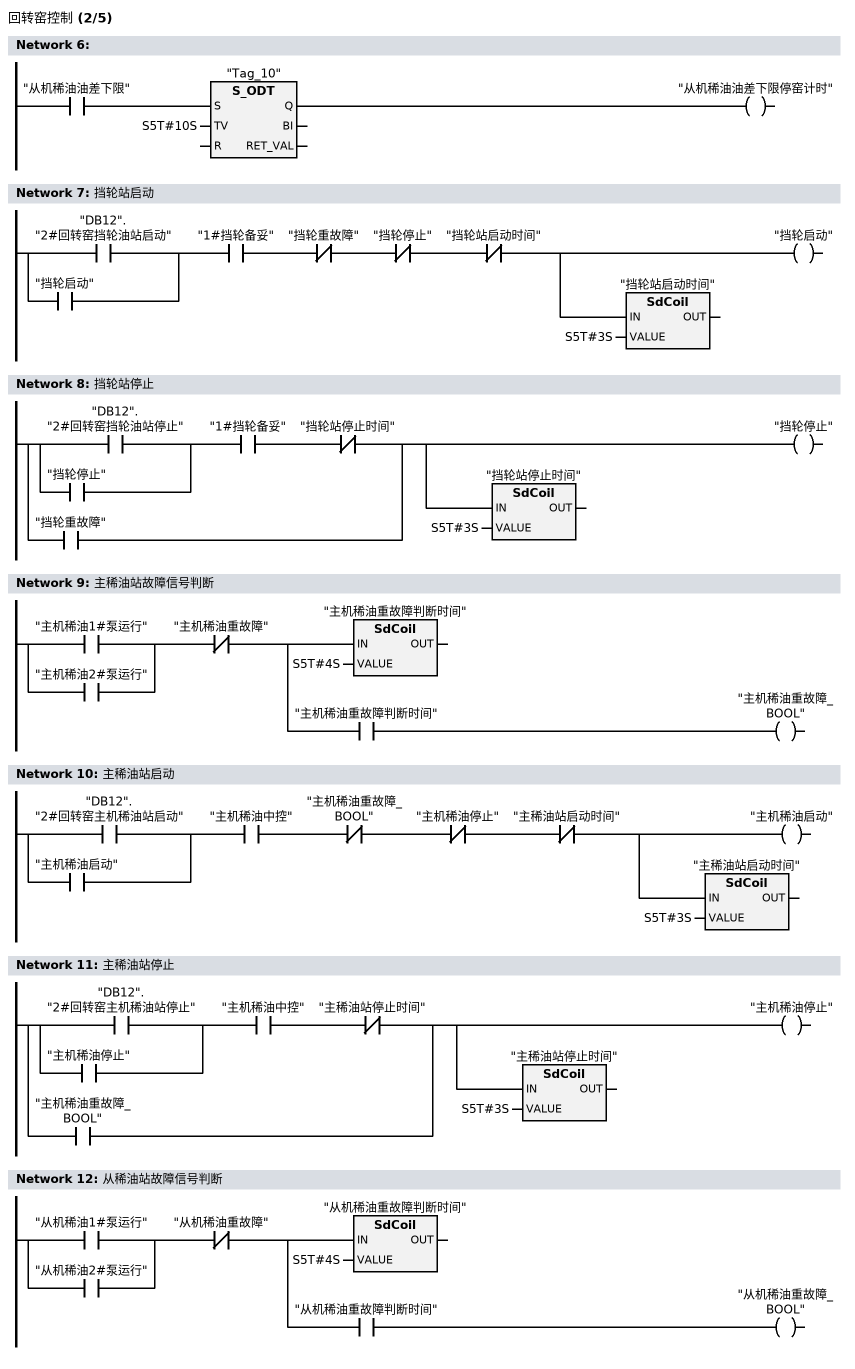
   RUNG wire#powerrail
      Contact( "从机稀油油差下限" )
      S_ODT(T_NO := "Tag_10", TV := S5T#10S, R :=, BI =>, RET_VAL =>)
      Coil( "从机稀油油差下限停窑计时" )
   END_RUNG
   // the same network as SCL:
   #_s5time1 := S_ODT(T_NO := "Tag_10", TV := S5T#10S, S := "从机稀油油差下限", Q => #_w1);
   "从机稀油油差下限停窑计时" := #_w1;
END_REGION

REGION Network 7: 挡轮站启动
   // no SCL statement known for SdCoil: written as a call
   "挡轮启动" := ("DB12"."2#回转窑挡轮油站启动" OR "挡轮启动") AND "1#挡轮备妥" AND NOT "挡轮重故障" AND NOT "挡轮停止" AND NOT "挡轮站启动时间";
   SdCoil(in := "挡轮启动", value := S5T#3S, operand := "挡轮站启动时间");
END_REGION

REGION Network 8: 挡轮站停止
   // no SCL statement known for SdCoil: written as a call
   "挡轮停止" := (("DB12"."2#回转窑挡轮油站停止" OR "挡轮停止") AND "1#挡轮备妥" AND NOT "挡轮站停止时间") OR "挡轮重故障";
   SdCoil(in := "挡轮停止", value := S5T#3S, operand := "挡轮站停止时间");
END_REGION

REGION Network 9: 主稀油站故障信号判断
   // no SCL statement known for SdCoil: written as a call
   #_w1 := ("主机稀油1#泵运行" OR "主机稀油2#泵运行") AND NOT "主机稀油重故障";
   SdCoil(in := #_w1, value := S5T#4S, operand := "主机稀油重故障判断时间");
   "主机稀油重故障_BOOL" := #_w1 AND "主机稀油重故障判断时间";
END_REGION

REGION Network 10: 主稀油站启动
   // no SCL statement known for SdCoil: written as a call
   "主机稀油启动" := ("DB12"."2#回转窑主机稀油站启动" OR "主机稀油启动") AND "主机稀油中控" AND NOT "主机稀油重故障_BOOL" AND NOT "主机稀油停止" AND NOT "主稀油站启动时间";
   SdCoil(in := "主机稀油启动", value := S5T#3S, operand := "主稀油站启动时间");
END_REGION

REGION Network 11: 主稀油站停止
   // no SCL statement known for SdCoil: written as a call
   "主机稀油停止" := (("DB12"."2#回转窑主机稀油站停止" OR "主机稀油停止") AND "主机稀油中控" AND NOT "主稀油站停止时间") OR "主机稀油重故障_BOOL";
   SdCoil(in := "主机稀油停止", value := S5T#3S, operand := "主稀油站停止时间");
END_REGION

REGION Network 12: 从稀油站故障信号判断
   // no SCL statement known for SdCoil: written as a call
   #_w1 := ("从机稀油1#泵运行" OR "从机稀油2#泵运行") AND NOT "从机稀油重故障";
   SdCoil(in := #_w1, value := S5T#4S, operand := "从机稀油重故障判断时间");
   "从机稀油重故障_BOOL" := #_w1 AND "从机稀油重故障判断时间";
END_REGION

REGION Network 13: 从稀油站启动
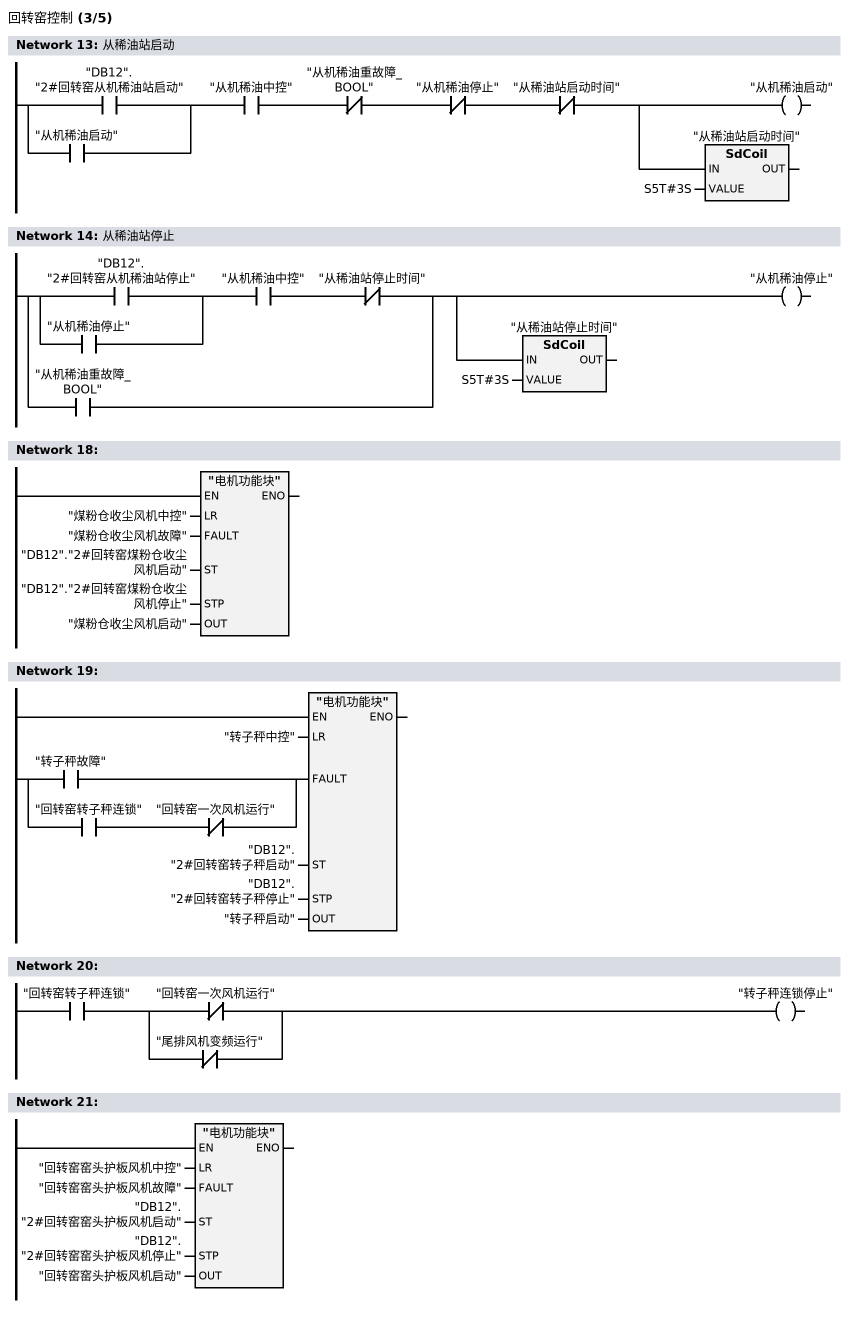
   // no SCL statement known for SdCoil: written as a call
   "从机稀油启动" := ("DB12"."2#回转窑从机稀油站启动" OR "从机稀油启动") AND "从机稀油中控" AND NOT "从机稀油重故障_BOOL" AND NOT "从机稀油停止" AND NOT "从稀油站启动时间";
   SdCoil(in := "从机稀油启动", value := S5T#3S, operand := "从稀油站启动时间");
END_REGION

REGION Network 14: 从稀油站停止
   // no SCL statement known for SdCoil: written as a call
   "从机稀油停止" := (("DB12"."2#回转窑从机稀油站停止" OR "从机稀油停止") AND "从机稀油中控" AND NOT "从稀油站停止时间") OR "从机稀油重故障_BOOL";
   SdCoil(in := "从机稀油停止", value := S5T#3S, operand := "从稀油站停止时间");
END_REGION

REGION Network 18
   RUNG wire#powerrail
      "电机功能块"(LR := "煤粉仓收尘风机中控", FAULT := "煤粉仓收尘风机故障", ST := "DB12"."2#回转窑煤粉仓收尘风机启动", STP := "DB12"."2#回转窑煤粉仓收尘风机停止", OUT := "煤粉仓收尘风机启动")
   END_RUNG
   // the same network as SCL:
   "电机功能块"(LR := "煤粉仓收尘风机中控",
           FAULT := "煤粉仓收尘风机故障",
           ST := "DB12"."2#回转窑煤粉仓收尘风机启动",
           STP := "DB12"."2#回转窑煤粉仓收尘风机停止",
           OUT := "煤粉仓收尘风机启动");
END_REGION

REGION Network 19
   RUNG wire#powerrail
      "电机功能块"(FAULT := wire#w1, LR := "转子秤中控", ST := "DB12"."2#回转窑转子秤启动", STP := "DB12"."2#回转窑转子秤停止", OUT := "转子秤启动")
   END_RUNG
   RUNG wire#powerrail
      Contact( "转子秤故障" )
   END_RUNG wire#w1
   RUNG wire#powerrail
      Contact( "回转窑转子秤连锁" )
      I_Contact( "回转窑一次风机运行" )
   END_RUNG wire#w1
   // the same network as SCL:
   "电机功能块"(LR := "转子秤中控",
           FAULT := "转子秤故障" OR ("回转窑转子秤连锁" AND NOT "回转窑一次风机运行"),
           ST := "DB12"."2#回转窑转子秤启动",
           STP := "DB12"."2#回转窑转子秤停止",
           OUT := "转子秤启动");
END_REGION

REGION Network 20
   RUNG wire#powerrail
      Contact( "回转窑转子秤连锁" )
      wire#w1
      I_Contact( "回转窑一次风机运行" )
      wire#w2
      Coil( "转子秤连锁停止" )
   END_RUNG
   RUNG wire#w1
      I_Contact( "尾排风机变频运行" )
   END_RUNG wire#w2
   // the same network as SCL:
   "转子秤连锁停止" := "回转窑转子秤连锁" AND (NOT "回转窑一次风机运行" OR NOT "尾排风机变频运行");
END_REGION

REGION Network 21
   RUNG wire#powerrail
      "电机功能块"(LR := "回转窑窑头护板风机中控", FAULT := "回转窑窑头护板风机故障", ST := "DB12"."2#回转窑窑头护板风机启动", STP := "DB12"."2#回转窑窑头护板风机停止", OUT := "回转窑窑头护板风机启动")
   END_RUNG
   // the same network as SCL:
   "电机功能块"(LR := "回转窑窑头护板风机中控",
           FAULT := "回转窑窑头护板风机故障",
           ST := "DB12"."2#回转窑窑头护板风机启动",
           STP := "DB12"."2#回转窑窑头护板风机停止",
           OUT := "回转窑窑头护板风机启动");
END_REGION

REGION Network 22
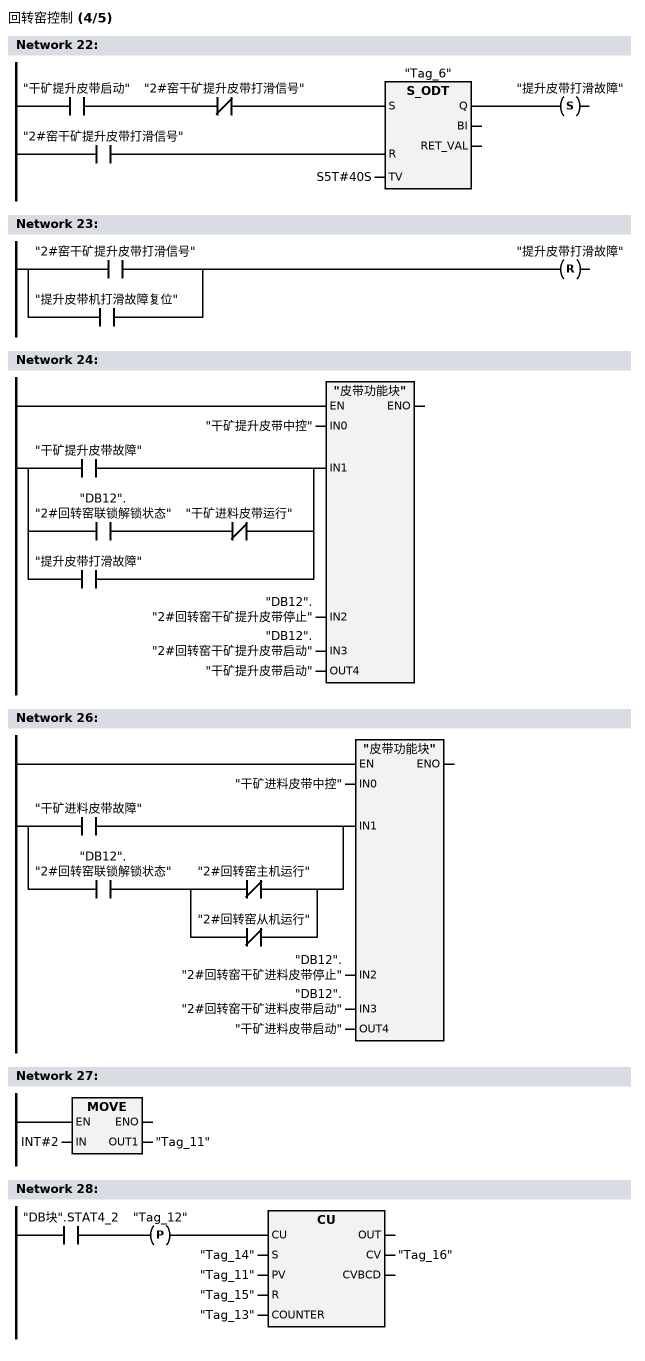
   RUNG wire#powerrail
      Contact( "干矿提升皮带启动" )
      I_Contact( "2#窑干矿提升皮带打滑信号" )
      S_ODT(T_NO := "Tag_6", R := wire#w1, TV := S5T#40S, BI =>, RET_VAL =>)
      S_Coil( "提升皮带打滑故障" )
   END_RUNG
   RUNG wire#powerrail
      Contact( "2#窑干矿提升皮带打滑信号" )
   END_RUNG wire#w1
   // the same network as SCL:
   #_s5time1 := S_ODT(T_NO := "Tag_6",
                      S := "干矿提升皮带启动" AND NOT "2#窑干矿提升皮带打滑信号",
                      R := "2#窑干矿提升皮带打滑信号",
                      TV := S5T#40S,
                      Q => #_w1);
   IF #_w1 THEN "提升皮带打滑故障" := TRUE; END_IF;
END_REGION

REGION Network 23
   RUNG wire#powerrail
      Contact( "2#窑干矿提升皮带打滑信号" )
      wire#w1
      R_Coil( "提升皮带打滑故障" )
   END_RUNG
   RUNG wire#powerrail
      Contact( "提升皮带机打滑故障复位" )
   END_RUNG wire#w1
   // the same network as SCL:
   IF "2#窑干矿提升皮带打滑信号" OR "提升皮带机打滑故障复位" THEN "提升皮带打滑故障" := FALSE; END_IF;
END_REGION

REGION Network 24
   RUNG wire#powerrail
      "皮带功能块"(IN1 := wire#w1, IN0 := "干矿提升皮带中控", IN2 := "DB12"."2#回转窑干矿提升皮带停止", IN3 := "DB12"."2#回转窑干矿提升皮带启动", OUT4 := "干矿提升皮带启动")
   END_RUNG
   RUNG wire#powerrail
      Contact( "干矿提升皮带故障" )
   END_RUNG wire#w1
   RUNG wire#powerrail
      Contact( "DB12"."2#回转窑联锁解锁状态" )
      I_Contact( "干矿进料皮带运行" )
   END_RUNG wire#w1
   RUNG wire#powerrail
      Contact( "提升皮带打滑故障" )
   END_RUNG wire#w1
   // the same network as SCL:
   "皮带功能块"(IN0 := "干矿提升皮带中控",
           IN1 := "干矿提升皮带故障" OR ("DB12"."2#回转窑联锁解锁状态" AND NOT "干矿进料皮带运行") OR "提升皮带打滑故障",
           IN2 := "DB12"."2#回转窑干矿提升皮带停止",
           IN3 := "DB12"."2#回转窑干矿提升皮带启动",
           OUT4 := "干矿提升皮带启动");
END_REGION

REGION Network 26
   RUNG wire#powerrail
      "皮带功能块"(IN1 := wire#w2, IN0 := "干矿进料皮带中控", IN2 := "DB12"."2#回转窑干矿进料皮带停止", IN3 := "DB12"."2#回转窑干矿进料皮带启动", OUT4 := "干矿进料皮带启动")
   END_RUNG
   RUNG wire#powerrail
      Contact( "干矿进料皮带故障" )
   END_RUNG wire#w2
   RUNG wire#powerrail
      Contact( "DB12"."2#回转窑联锁解锁状态" )
      wire#w1
      I_Contact( "2#回转窑主机运行" )
   END_RUNG wire#w2
   RUNG wire#w1
      I_Contact( "2#回转窑从机运行" )
   END_RUNG wire#w2
   // the same network as SCL:
   "皮带功能块"(IN0 := "干矿进料皮带中控",
           IN1 := "干矿进料皮带故障" OR ("DB12"."2#回转窑联锁解锁状态" AND (NOT "2#回转窑主机运行" OR NOT "2#回转窑从机运行")),
           IN2 := "DB12"."2#回转窑干矿进料皮带停止",
           IN3 := "DB12"."2#回转窑干矿进料皮带启动",
           OUT4 := "干矿进料皮带启动");
END_REGION

REGION Network 27
   RUNG wire#powerrail
      { S7_GenerateENO := "TRUE" } Move(in := INT#2, out1 => "Tag_11")
   END_RUNG
   // the same network as SCL:
   "Tag_11" := INT#2;
END_REGION

REGION Network 28
   // no SCL statement known for Cu: written as a call
   #_w1 := "DB块".STAT4_2 AND NOT "Tag_12";   // rising edge
   "Tag_12" := "DB块".STAT4_2;
   Cu(cu := #_w1, s := "Tag_14", pv := "Tag_11", r := "Tag_15", "counter" := "Tag_13", cv => "Tag_16");
END_REGION

REGION Network 29
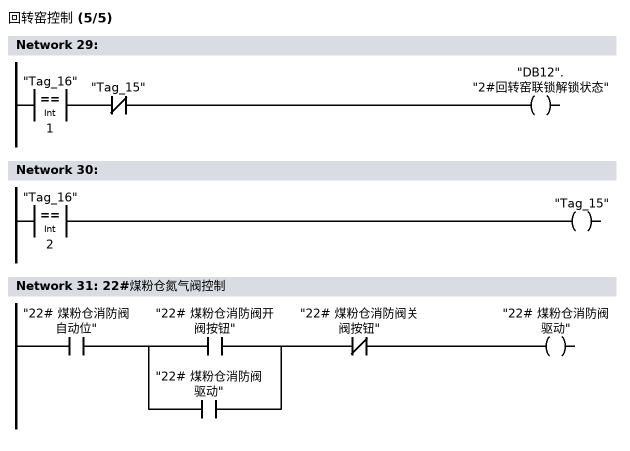
   RUNG wire#powerrail
      { S7_Templates := "SrcType := Int" } EQ_Contact(in1 := "Tag_16", in2 := 1)
      I_Contact( "Tag_15" )
      Coil( "DB12"."2#回转窑联锁解锁状态" )
   END_RUNG
   // the same network as SCL:
   "DB12"."2#回转窑联锁解锁状态" := ("Tag_16" = 1) AND NOT "Tag_15";
END_REGION

REGION Network 30
   RUNG wire#powerrail
      { S7_Templates := "SrcType := Int" } EQ_Contact(in1 := "Tag_16", in2 := 2)
      Coil( "Tag_15" )
   END_RUNG
   // the same network as SCL:
   "Tag_15" := "Tag_16" = 2;
END_REGION

REGION Network 31: 22#煤粉仓氮气阀控制
   RUNG wire#powerrail
      Contact( "22# 煤粉仓消防阀自动位" )
      wire#w1
      Contact( "22# 煤粉仓消防阀开阀按钮" )
      wire#w2
      I_Contact( "22# 煤粉仓消防阀关阀按钮" )
      Coil( "22# 煤粉仓消防阀驱动" )
   END_RUNG
   RUNG wire#w1
      Contact( "22# 煤粉仓消防阀驱动" )
   END_RUNG wire#w2
   // the same network as SCL:
   "22# 煤粉仓消防阀驱动" := "22# 煤粉仓消防阀自动位" AND ("22# 煤粉仓消防阀开阀按钮" OR "22# 煤粉仓消防阀驱动") AND NOT "22# 煤粉仓消防阀关阀按钮";
END_REGION
END_FUNCTION

FUNCTION "回转窑模拟量反馈" : Void   // FC12, LAD
{ S7_Optimized_Access := 'FALSE' }
VERSION : 0.1
   VAR_TEMP   // added for the SCL form of the ladder/FBD networks
      _w1 : Bool;
      _s5time1 : S5Time;
   END_VAR
BEGIN

REGION Network 1
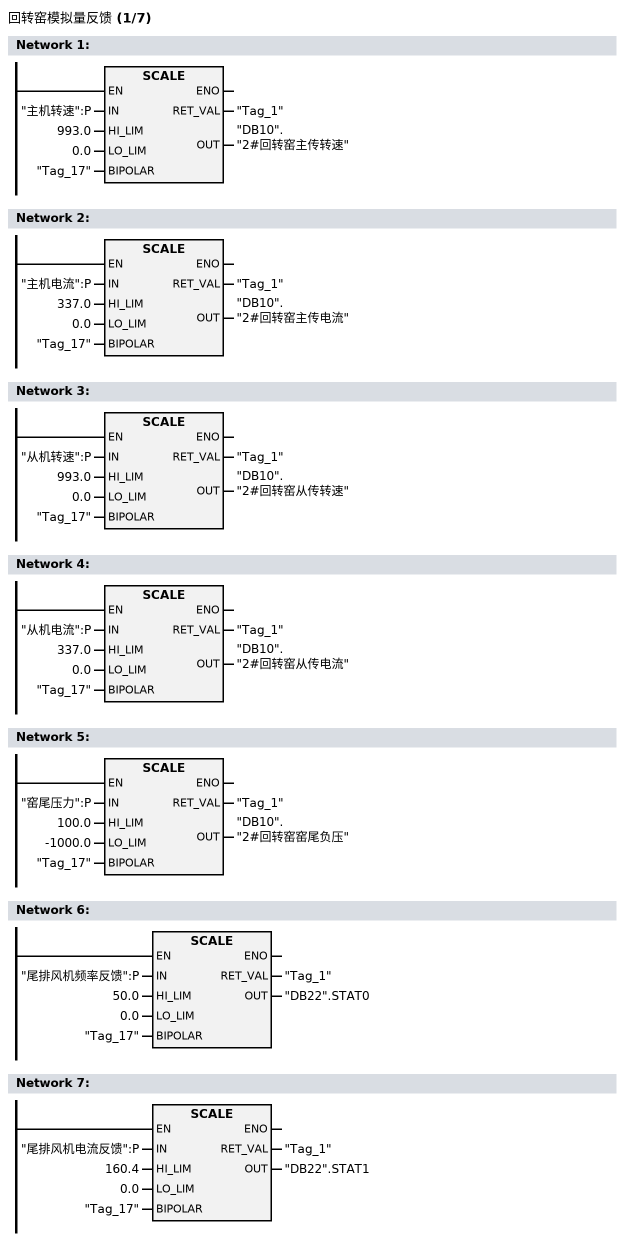
   "Tag_1" := SCALE(IN := "主机转速":P,
                    HI_LIM := 993.0,
                    LO_LIM := 0.0,
                    BIPOLAR := "Tag_17",
                    OUT => "DB10"."2#回转窑主传转速");
END_REGION

REGION Network 2
   "Tag_1" := SCALE(IN := "主机电流":P,
                    HI_LIM := 337.0,
                    LO_LIM := 0.0,
                    BIPOLAR := "Tag_17",
                    OUT => "DB10"."2#回转窑主传电流");
END_REGION

REGION Network 3
   "Tag_1" := SCALE(IN := "从机转速":P,
                    HI_LIM := 993.0,
                    LO_LIM := 0.0,
                    BIPOLAR := "Tag_17",
                    OUT => "DB10"."2#回转窑从传转速");
END_REGION

REGION Network 4
   "Tag_1" := SCALE(IN := "从机电流":P,
                    HI_LIM := 337.0,
                    LO_LIM := 0.0,
                    BIPOLAR := "Tag_17",
                    OUT => "DB10"."2#回转窑从传电流");
END_REGION

REGION Network 5
   "Tag_1" := SCALE(IN := "窑尾压力":P,
                    HI_LIM := 100.0,
                    LO_LIM := -1000.0,
                    BIPOLAR := "Tag_17",
                    OUT => "DB10"."2#回转窑窑尾负压");
END_REGION

REGION Network 6
   "Tag_1" := SCALE(IN := "尾排风机频率反馈":P, HI_LIM := 50.0, LO_LIM := 0.0, BIPOLAR := "Tag_17", OUT => "DB22".STAT0);
END_REGION

REGION Network 7
   "Tag_1" := SCALE(IN := "尾排风机电流反馈":P,
                    HI_LIM := 160.4,
                    LO_LIM := 0.0,
                    BIPOLAR := "Tag_17",
                    OUT => "DB22".STAT1);
END_REGION

REGION Network 8
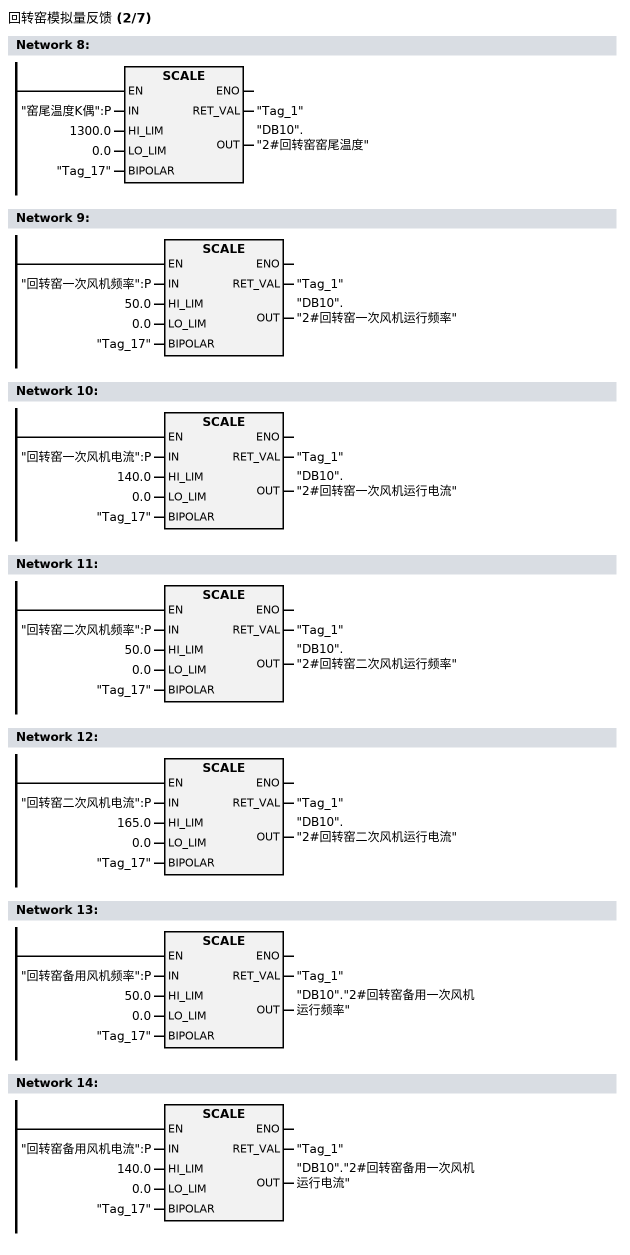
   "Tag_1" := SCALE(IN := "窑尾温度K偶":P,
                    HI_LIM := 1300.0,
                    LO_LIM := 0.0,
                    BIPOLAR := "Tag_17",
                    OUT => "DB10"."2#回转窑窑尾温度");
END_REGION

REGION Network 9
   "Tag_1" := SCALE(IN := "回转窑一次风机频率":P,
                    HI_LIM := 50.0,
                    LO_LIM := 0.0,
                    BIPOLAR := "Tag_17",
                    OUT => "DB10"."2#回转窑一次风机运行频率");
END_REGION

REGION Network 10
   "Tag_1" := SCALE(IN := "回转窑一次风机电流":P,
                    HI_LIM := 140.0,
                    LO_LIM := 0.0,
                    BIPOLAR := "Tag_17",
                    OUT => "DB10"."2#回转窑一次风机运行电流");
END_REGION

REGION Network 11
   "Tag_1" := SCALE(IN := "回转窑二次风机频率":P,
                    HI_LIM := 50.0,
                    LO_LIM := 0.0,
                    BIPOLAR := "Tag_17",
                    OUT => "DB10"."2#回转窑二次风机运行频率");
END_REGION

REGION Network 12
   "Tag_1" := SCALE(IN := "回转窑二次风机电流":P,
                    HI_LIM := 165.0,
                    LO_LIM := 0.0,
                    BIPOLAR := "Tag_17",
                    OUT => "DB10"."2#回转窑二次风机运行电流");
END_REGION

REGION Network 13
   "Tag_1" := SCALE(IN := "回转窑备用风机频率":P,
                    HI_LIM := 50.0,
                    LO_LIM := 0.0,
                    BIPOLAR := "Tag_17",
                    OUT => "DB10"."2#回转窑备用一次风机运行频率");
END_REGION

REGION Network 14
   "Tag_1" := SCALE(IN := "回转窑备用风机电流":P,
                    HI_LIM := 140.0,
                    LO_LIM := 0.0,
                    BIPOLAR := "Tag_17",
                    OUT => "DB10"."2#回转窑备用一次风机运行电流");
END_REGION

REGION Network 15
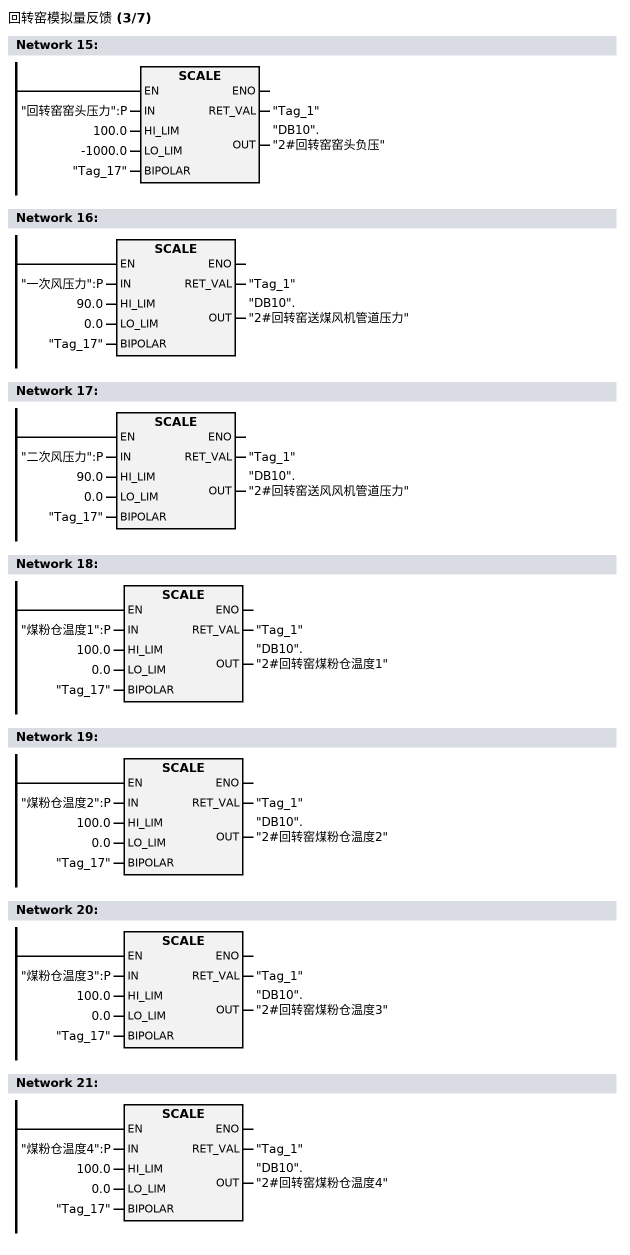
   "Tag_1" := SCALE(IN := "回转窑窑头压力":P,
                    HI_LIM := 100.0,
                    LO_LIM := -1000.0,
                    BIPOLAR := "Tag_17",
                    OUT => "DB10"."2#回转窑窑头负压");
END_REGION

REGION Network 16
   "Tag_1" := SCALE(IN := "一次风压力":P,
                    HI_LIM := 90.0,
                    LO_LIM := 0.0,
                    BIPOLAR := "Tag_17",
                    OUT => "DB10"."2#回转窑送煤风机管道压力");
END_REGION

REGION Network 17
   "Tag_1" := SCALE(IN := "二次风压力":P,
                    HI_LIM := 90.0,
                    LO_LIM := 0.0,
                    BIPOLAR := "Tag_17",
                    OUT => "DB10"."2#回转窑送风风机管道压力");
END_REGION

REGION Network 18
   "Tag_1" := SCALE(IN := "煤粉仓温度1":P,
                    HI_LIM := 100.0,
                    LO_LIM := 0.0,
                    BIPOLAR := "Tag_17",
                    OUT => "DB10"."2#回转窑煤粉仓温度1");
END_REGION

REGION Network 19
   "Tag_1" := SCALE(IN := "煤粉仓温度2":P,
                    HI_LIM := 100.0,
                    LO_LIM := 0.0,
                    BIPOLAR := "Tag_17",
                    OUT => "DB10"."2#回转窑煤粉仓温度2");
END_REGION

REGION Network 20
   "Tag_1" := SCALE(IN := "煤粉仓温度3":P,
                    HI_LIM := 100.0,
                    LO_LIM := 0.0,
                    BIPOLAR := "Tag_17",
                    OUT => "DB10"."2#回转窑煤粉仓温度3");
END_REGION

REGION Network 21
   "Tag_1" := SCALE(IN := "煤粉仓温度4":P,
                    HI_LIM := 100.0,
                    LO_LIM := 0.0,
                    BIPOLAR := "Tag_17",
                    OUT => "DB10"."2#回转窑煤粉仓温度4");
END_REGION

REGION Network 22
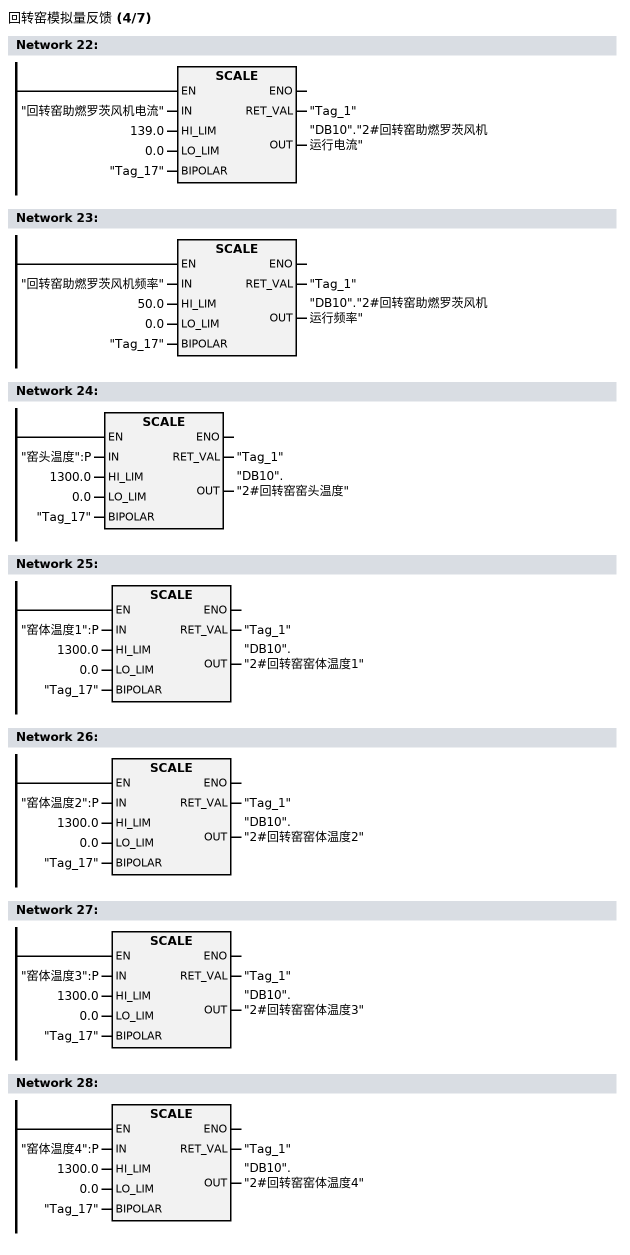
   "Tag_1" := SCALE(IN := "回转窑助燃罗茨风机电流",
                    HI_LIM := 139.0,
                    LO_LIM := 0.0,
                    BIPOLAR := "Tag_17",
                    OUT => "DB10"."2#回转窑助燃罗茨风机运行电流");
END_REGION

REGION Network 23
   "Tag_1" := SCALE(IN := "回转窑助燃罗茨风机频率",
                    HI_LIM := 50.0,
                    LO_LIM := 0.0,
                    BIPOLAR := "Tag_17",
                    OUT => "DB10"."2#回转窑助燃罗茨风机运行频率");
END_REGION

REGION Network 24
   "Tag_1" := SCALE(IN := "窑头温度":P,
                    HI_LIM := 1300.0,
                    LO_LIM := 0.0,
                    BIPOLAR := "Tag_17",
                    OUT => "DB10"."2#回转窑窑头温度");
END_REGION

REGION Network 25
   "Tag_1" := SCALE(IN := "窑体温度1":P,
                    HI_LIM := 1300.0,
                    LO_LIM := 0.0,
                    BIPOLAR := "Tag_17",
                    OUT => "DB10"."2#回转窑窑体温度1");
END_REGION

REGION Network 26
   "Tag_1" := SCALE(IN := "窑体温度2":P,
                    HI_LIM := 1300.0,
                    LO_LIM := 0.0,
                    BIPOLAR := "Tag_17",
                    OUT => "DB10"."2#回转窑窑体温度2");
END_REGION

REGION Network 27
   "Tag_1" := SCALE(IN := "窑体温度3":P,
                    HI_LIM := 1300.0,
                    LO_LIM := 0.0,
                    BIPOLAR := "Tag_17",
                    OUT => "DB10"."2#回转窑窑体温度3");
END_REGION

REGION Network 28
   "Tag_1" := SCALE(IN := "窑体温度4":P,
                    HI_LIM := 1300.0,
                    LO_LIM := 0.0,
                    BIPOLAR := "Tag_17",
                    OUT => "DB10"."2#回转窑窑体温度4");
END_REGION

REGION Network 29
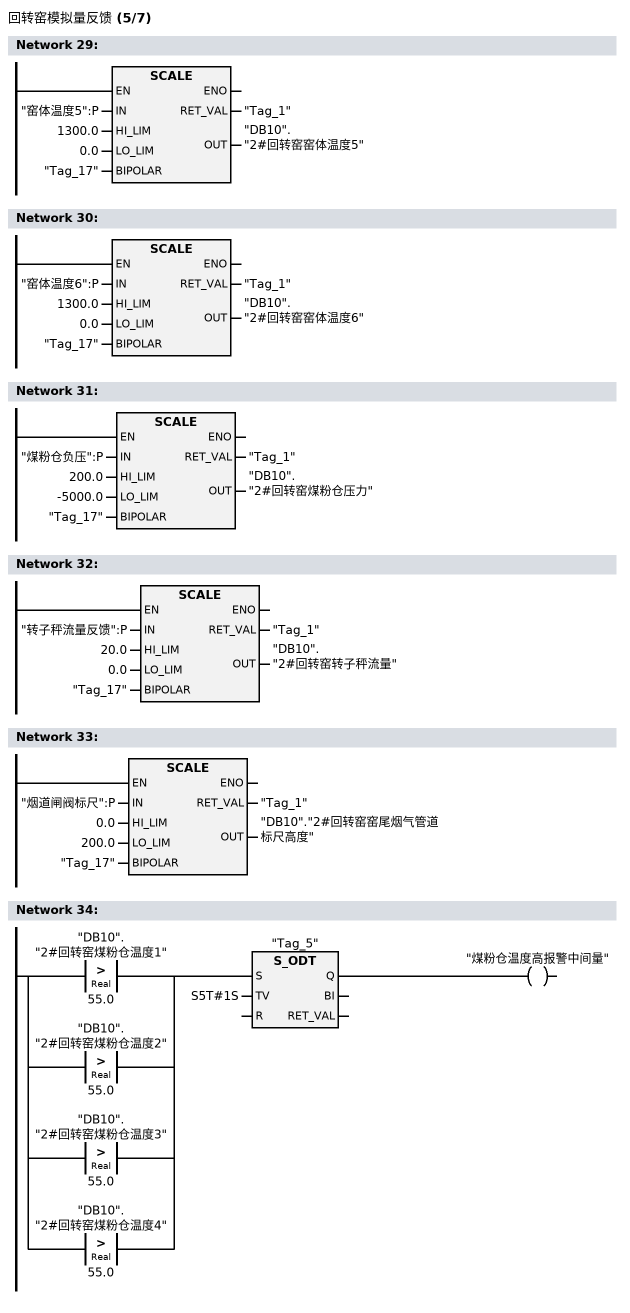
   "Tag_1" := SCALE(IN := "窑体温度5":P,
                    HI_LIM := 1300.0,
                    LO_LIM := 0.0,
                    BIPOLAR := "Tag_17",
                    OUT => "DB10"."2#回转窑窑体温度5");
END_REGION

REGION Network 30
   "Tag_1" := SCALE(IN := "窑体温度6":P,
                    HI_LIM := 1300.0,
                    LO_LIM := 0.0,
                    BIPOLAR := "Tag_17",
                    OUT => "DB10"."2#回转窑窑体温度6");
END_REGION

REGION Network 31
   "Tag_1" := SCALE(IN := "煤粉仓负压":P,
                    HI_LIM := 200.0,
                    LO_LIM := -5000.0,
                    BIPOLAR := "Tag_17",
                    OUT => "DB10"."2#回转窑煤粉仓压力");
END_REGION

REGION Network 32
   "Tag_1" := SCALE(IN := "转子秤流量反馈":P,
                    HI_LIM := 20.0,
                    LO_LIM := 0.0,
                    BIPOLAR := "Tag_17",
                    OUT => "DB10"."2#回转窑转子秤流量");
END_REGION

REGION Network 33
   "Tag_1" := SCALE(IN := "烟道闸阀标尺":P,
                    HI_LIM := 0.0,
                    LO_LIM := 200.0,
                    BIPOLAR := "Tag_17",
                    OUT => "DB10"."2#回转窑窑尾烟气管道标尺高度");
END_REGION

REGION Network 34
   RUNG wire#powerrail
      { S7_Templates := "SrcType := Real" } GT_Contact(in1 := "DB10"."2#回转窑煤粉仓温度1", in2 := 55.0)
      wire#w1
      S_ODT(T_NO := "Tag_5", TV := S5T#1S, R :=, BI =>, RET_VAL =>)
      Coil( "煤粉仓温度高报警中间量" )
   END_RUNG
   RUNG wire#powerrail
      { S7_Templates := "SrcType := Real" } GT_Contact(in1 := "DB10"."2#回转窑煤粉仓温度2", in2 := 55.0)
   END_RUNG wire#w1
   RUNG wire#powerrail
      { S7_Templates := "SrcType := Real" } GT_Contact(in1 := "DB10"."2#回转窑煤粉仓温度3", in2 := 55.0)
   END_RUNG wire#w1
   RUNG wire#powerrail
      { S7_Templates := "SrcType := Real" } GT_Contact(in1 := "DB10"."2#回转窑煤粉仓温度4", in2 := 55.0)
   END_RUNG wire#w1
   // the same network as SCL:
   #_s5time1 := S_ODT(T_NO := "Tag_5",
                      S := ("DB10"."2#回转窑煤粉仓温度1" > 55.0) OR ("DB10"."2#回转窑煤粉仓温度2" > 55.0) OR ("DB10"."2#回转窑煤粉仓温度3" > 55.0) OR ("DB10"."2#回转窑煤粉仓温度4" > 55.0),
                      TV := S5T#1S,
                      Q => #_w1);
   "煤粉仓温度高报警中间量" := #_w1;
END_REGION

REGION Network 35
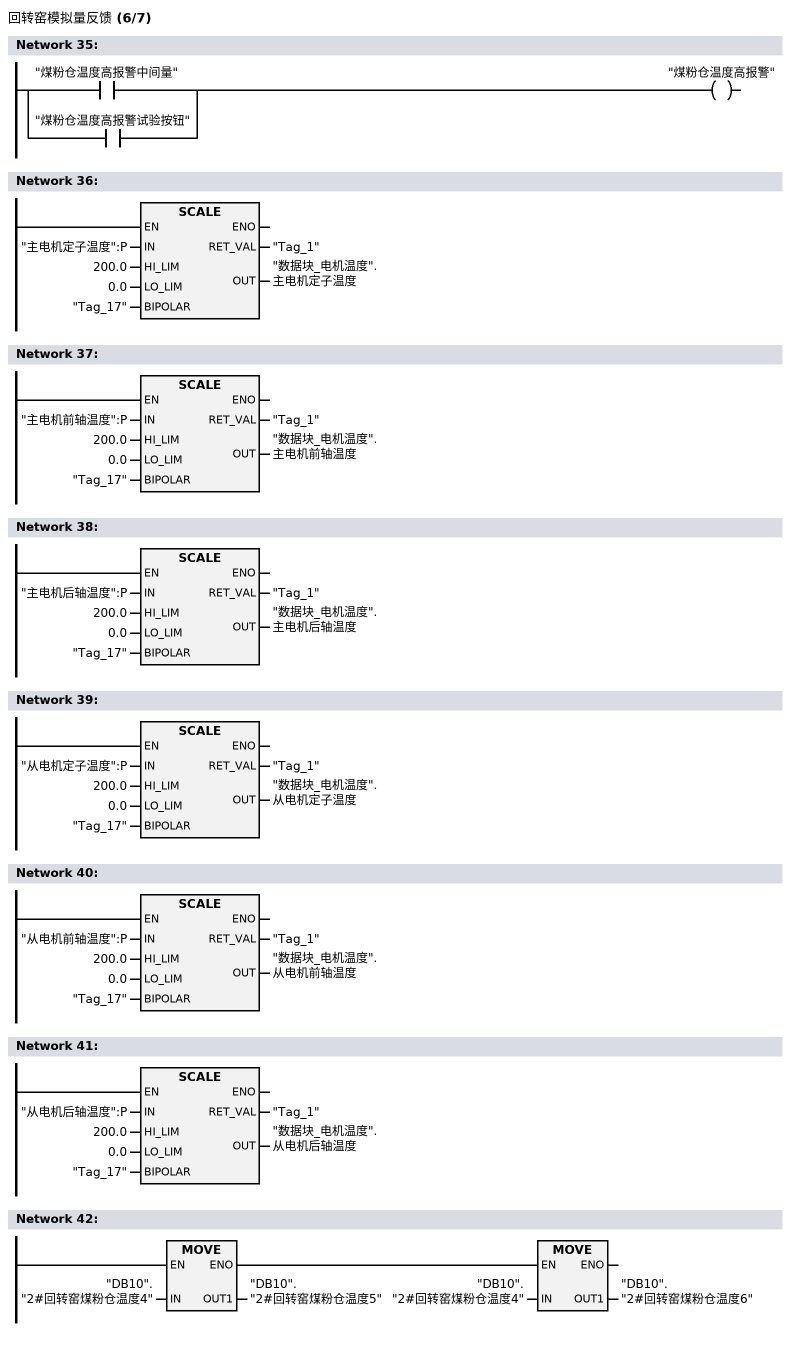
   RUNG wire#powerrail
      Contact( "煤粉仓温度高报警中间量" )
      wire#w1
      Coil( "煤粉仓温度高报警" )
   END_RUNG
   RUNG wire#powerrail
      Contact( "煤粉仓温度高报警试验按钮" )
   END_RUNG wire#w1
   // the same network as SCL:
   "煤粉仓温度高报警" := "煤粉仓温度高报警中间量" OR "煤粉仓温度高报警试验按钮";
END_REGION

REGION Network 36
   "Tag_1" := SCALE(IN := "主电机定子温度":P,
                    HI_LIM := 200.0,
                    LO_LIM := 0.0,
                    BIPOLAR := "Tag_17",
                    OUT => "数据块_电机温度".主电机定子温度);
END_REGION

REGION Network 37
   "Tag_1" := SCALE(IN := "主电机前轴温度":P,
                    HI_LIM := 200.0,
                    LO_LIM := 0.0,
                    BIPOLAR := "Tag_17",
                    OUT => "数据块_电机温度".主电机前轴温度);
END_REGION

REGION Network 38
   "Tag_1" := SCALE(IN := "主电机后轴温度":P,
                    HI_LIM := 200.0,
                    LO_LIM := 0.0,
                    BIPOLAR := "Tag_17",
                    OUT => "数据块_电机温度".主电机后轴温度);
END_REGION

REGION Network 39
   "Tag_1" := SCALE(IN := "从电机定子温度":P,
                    HI_LIM := 200.0,
                    LO_LIM := 0.0,
                    BIPOLAR := "Tag_17",
                    OUT => "数据块_电机温度".从电机定子温度);
END_REGION

REGION Network 40
   "Tag_1" := SCALE(IN := "从电机前轴温度":P,
                    HI_LIM := 200.0,
                    LO_LIM := 0.0,
                    BIPOLAR := "Tag_17",
                    OUT => "数据块_电机温度".从电机前轴温度);
END_REGION

REGION Network 41
   "Tag_1" := SCALE(IN := "从电机后轴温度":P,
                    HI_LIM := 200.0,
                    LO_LIM := 0.0,
                    BIPOLAR := "Tag_17",
                    OUT => "数据块_电机温度".从电机后轴温度);
END_REGION

REGION Network 42
   RUNG wire#powerrail
      Move(in := "DB10"."2#回转窑煤粉仓温度4", out1 => "DB10"."2#回转窑煤粉仓温度5")
      Move(in := "DB10"."2#回转窑煤粉仓温度4", out1 => "DB10"."2#回转窑煤粉仓温度6")
   END_RUNG
   // the same network as SCL:
   "DB10"."2#回转窑煤粉仓温度5" := "DB10"."2#回转窑煤粉仓温度4";
   "DB10"."2#回转窑煤粉仓温度6" := "DB10"."2#回转窑煤粉仓温度4";
END_REGION

REGION Network 43: 2#回转窑富氧流量
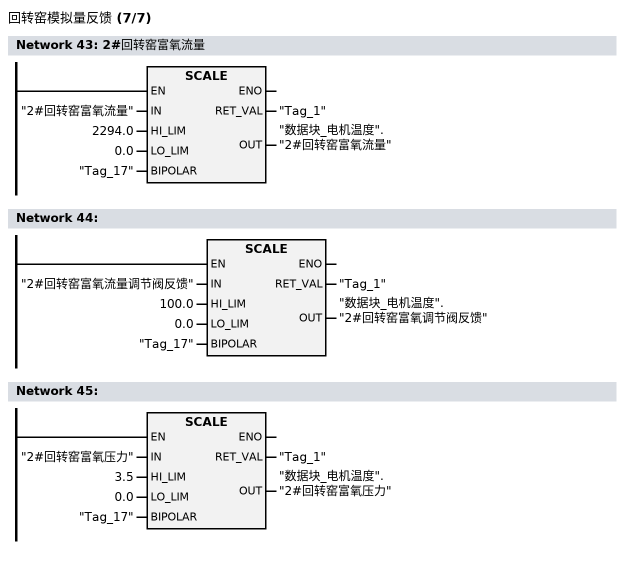
   "Tag_1" := SCALE(IN := "2#回转窑富氧流量",
                    HI_LIM := 2294.0,
                    LO_LIM := 0.0,
                    BIPOLAR := "Tag_17",
                    OUT => "数据块_电机温度"."2#回转窑富氧流量");
END_REGION

REGION Network 44
   "Tag_1" := SCALE(IN := "2#回转窑富氧流量调节阀反馈",
                    HI_LIM := 100.0,
                    LO_LIM := 0.0,
                    BIPOLAR := "Tag_17",
                    OUT => "数据块_电机温度"."2#回转窑富氧调节阀反馈");
END_REGION

REGION Network 45
   "Tag_1" := SCALE(IN := "2#回转窑富氧压力",
                    HI_LIM := 3.5,
                    LO_LIM := 0.0,
                    BIPOLAR := "Tag_17",
                    OUT => "数据块_电机温度"."2#回转窑富氧压力");
END_REGION
END_FUNCTION

FUNCTION "回转窑风机控制" : Void   // FC13, LAD
{ S7_Optimized_Access := 'FALSE' }
VERSION : 0.1
   VAR_TEMP   // added for the SCL form of the ladder/FBD networks
      _w1 : Bool;
      _s5time1 : S5Time;
   END_VAR
BEGIN

REGION Network 1
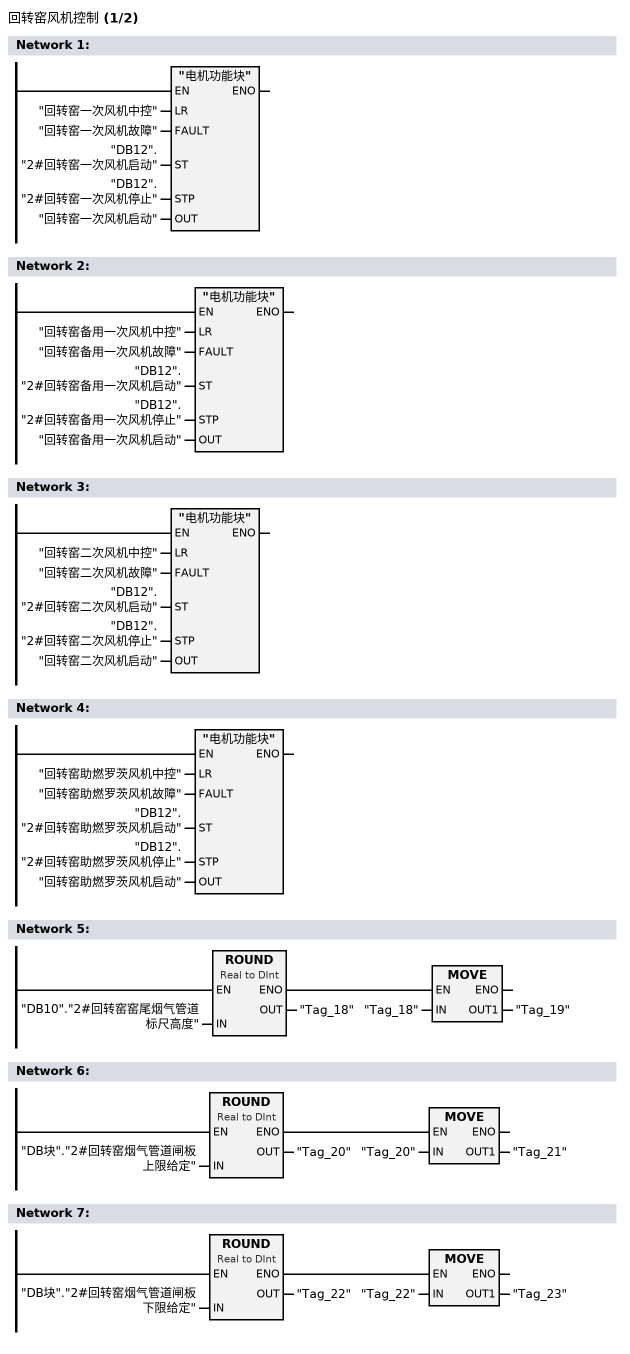
   RUNG wire#powerrail
      "电机功能块"(LR := "回转窑一次风机中控", FAULT := "回转窑一次风机故障", ST := "DB12"."2#回转窑一次风机启动", STP := "DB12"."2#回转窑一次风机停止", OUT := "回转窑一次风机启动")
   END_RUNG
   // the same network as SCL:
   "电机功能块"(LR := "回转窑一次风机中控",
           FAULT := "回转窑一次风机故障",
           ST := "DB12"."2#回转窑一次风机启动",
           STP := "DB12"."2#回转窑一次风机停止",
           OUT := "回转窑一次风机启动");
END_REGION

REGION Network 2
   RUNG wire#powerrail
      "电机功能块"(LR := "回转窑备用一次风机中控", FAULT := "回转窑备用一次风机故障", ST := "DB12"."2#回转窑备用一次风机启动", STP := "DB12"."2#回转窑备用一次风机停止", OUT := "回转窑备用一次风机启动")
   END_RUNG
   // the same network as SCL:
   "电机功能块"(LR := "回转窑备用一次风机中控",
           FAULT := "回转窑备用一次风机故障",
           ST := "DB12"."2#回转窑备用一次风机启动",
           STP := "DB12"."2#回转窑备用一次风机停止",
           OUT := "回转窑备用一次风机启动");
END_REGION

REGION Network 3
   RUNG wire#powerrail
      "电机功能块"(LR := "回转窑二次风机中控", FAULT := "回转窑二次风机故障", ST := "DB12"."2#回转窑二次风机启动", STP := "DB12"."2#回转窑二次风机停止", OUT := "回转窑二次风机启动")
   END_RUNG
   // the same network as SCL:
   "电机功能块"(LR := "回转窑二次风机中控",
           FAULT := "回转窑二次风机故障",
           ST := "DB12"."2#回转窑二次风机启动",
           STP := "DB12"."2#回转窑二次风机停止",
           OUT := "回转窑二次风机启动");
END_REGION

REGION Network 4
   RUNG wire#powerrail
      "电机功能块"(LR := "回转窑助燃罗茨风机中控", FAULT := "回转窑助燃罗茨风机故障", ST := "DB12"."2#回转窑助燃罗茨风机启动", STP := "DB12"."2#回转窑助燃罗茨风机停止", OUT := "回转窑助燃罗茨风机启动")
   END_RUNG
   // the same network as SCL:
   "电机功能块"(LR := "回转窑助燃罗茨风机中控",
           FAULT := "回转窑助燃罗茨风机故障",
           ST := "DB12"."2#回转窑助燃罗茨风机启动",
           STP := "DB12"."2#回转窑助燃罗茨风机停止",
           OUT := "回转窑助燃罗茨风机启动");
END_REGION

REGION Network 5
   RUNG wire#powerrail
      { S7_Templates := "[SrcType := Real, DestType := DInt]"; S7_GenerateENO := "TRUE" } Round(in := "DB10"."2#回转窑窑尾烟气管道标尺高度", out => "Tag_18")
      { S7_GenerateENO := "TRUE" } Move(in := "Tag_18", out1 => "Tag_19")
   END_RUNG
   // the same network as SCL:
   // ENO of a box is taken as its EN; it also drops when the box reports an error
   "Tag_18" := ROUND("DB10"."2#回转窑窑尾烟气管道标尺高度");
   "Tag_19" := "Tag_18";
END_REGION

REGION Network 6
   RUNG wire#powerrail
      { S7_Templates := "[SrcType := Real, DestType := DInt]"; S7_GenerateENO := "TRUE" } Round(in := "DB块"."2#回转窑烟气管道闸板上限给定", out => "Tag_20")
      { S7_GenerateENO := "TRUE" } Move(in := "Tag_20", out1 => "Tag_21")
   END_RUNG
   // the same network as SCL:
   // ENO of a box is taken as its EN; it also drops when the box reports an error
   "Tag_20" := ROUND("DB块"."2#回转窑烟气管道闸板上限给定");
   "Tag_21" := "Tag_20";
END_REGION

REGION Network 7
   RUNG wire#powerrail
      { S7_Templates := "[SrcType := Real, DestType := DInt]"; S7_GenerateENO := "TRUE" } Round(in := "DB块"."2#回转窑烟气管道闸板下限给定", out => "Tag_22")
      { S7_GenerateENO := "TRUE" } Move(in := "Tag_22", out1 => "Tag_23")
   END_RUNG
   // the same network as SCL:
   // ENO of a box is taken as its EN; it also drops when the box reports an error
   "Tag_22" := ROUND("DB块"."2#回转窑烟气管道闸板下限给定");
   "Tag_23" := "Tag_22";
END_REGION

REGION Network 8
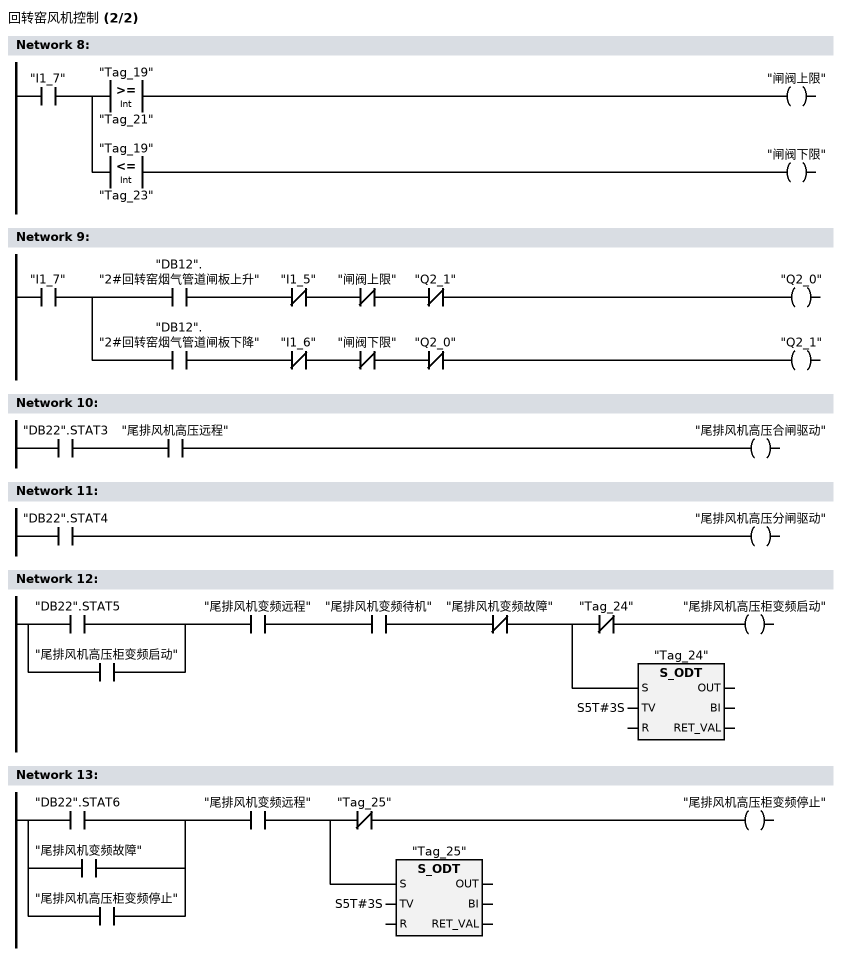
   RUNG wire#powerrail
      Contact( "I1_7" )
      wire#w1
      { S7_Templates := "SrcType := Int" } GE_Contact(in1 := "Tag_19", in2 := "Tag_21")
      Coil( "闸阀上限" )
   END_RUNG
   RUNG wire#w1
      { S7_Templates := "SrcType := Int" } LE_Contact(in1 := "Tag_19", in2 := "Tag_23")
      Coil( "闸阀下限" )
   END_RUNG
   // the same network as SCL:
   "闸阀上限" := "I1_7" AND ("Tag_19" >= "Tag_21");
   "闸阀下限" := "I1_7" AND ("Tag_19" <= "Tag_23");
END_REGION
